   "TT426_5S_ALM_ANALOG_DB_VERY HIGH LEVEL VALUE (HH)" : Real = PLC TT426_5S_ALM_ANALOG_DB."VERY HIGH LEVEL VALUE (HH)" AT %DB2082.DBD34, 1 s
   "TT426_5S_ALM_ANALOG_DB_VERY LOW LEVEL VALUE (LL)" : Real = PLC TT426_5S_ALM_ANALOG_DB."VERY LOW LEVEL VALUE (LL)" AT %DB2082.DBD22, 1 s
   "TT426_6P_ALM_ANALOG_DB_HIGH LEVEL VALUE (H)" : Real = PLC TT426_6P_ALM_ANALOG_DB."HIGH LEVEL VALUE (H)" AT %DB2083.DBD30, 1 s
   "TT426_6P_ALM_ANALOG_DB_LOW LEVEL VALUE (L)" : Real = PLC TT426_6P_ALM_ANALOG_DB."LOW LEVEL VALUE (L)" AT %DB2083.DBD26, 1 s
   "TT426_6P_ALM_ANALOG_DB_VERY HIGH LEVEL VALUE (HH)" : Real = PLC TT426_6P_ALM_ANALOG_DB."VERY HIGH LEVEL VALUE (HH)" AT %DB2083.DBD34, 1 s
   "TT426_6P_ALM_ANALOG_DB_VERY LOW LEVEL VALUE (LL)" : Real = PLC TT426_6P_ALM_ANALOG_DB."VERY LOW LEVEL VALUE (LL)" AT %DB2083.DBD22, 1 s
   "TT426_6S_ALM_ANALOG_DB_HIGH LEVEL VALUE (H)" : Real = PLC TT426_6S_ALM_ANALOG_DB."HIGH LEVEL VALUE (H)" AT %DB2085.DBD30, 1 s
   "TT426_6S_ALM_ANALOG_DB_LOW LEVEL VALUE (L)" : Real = PLC TT426_6S_ALM_ANALOG_DB."LOW LEVEL VALUE (L)" AT %DB2085.DBD26, 1 s
   "TT426_6S_ALM_ANALOG_DB_VERY HIGH LEVEL VALUE (HH)" : Real = PLC TT426_6S_ALM_ANALOG_DB."VERY HIGH LEVEL VALUE (HH)" AT %DB2085.DBD34, 1 s
   "TT426_6S_ALM_ANALOG_DB_VERY LOW LEVEL VALUE (LL)" : Real = PLC TT426_6S_ALM_ANALOG_DB."VERY LOW LEVEL VALUE (LL)" AT %DB2085.DBD22, 1 s
   "TT426_APT_ALM_ANALOG_DB_HIGH LEVEL VALUE (H)" : Real = PLC TT426_APT_ALM_ANALOG_DB."HIGH LEVEL VALUE (H)" AT %DB2087.DBD30, 1 s
   "TT426_APT_ALM_ANALOG_DB_LOW LEVEL VALUE (L)" : Real = PLC TT426_APT_ALM_ANALOG_DB."LOW LEVEL VALUE (L)" AT %DB2087.DBD26, 1 s
   "TT426_APT_ALM_ANALOG_DB_VERY HIGH LEVEL VALUE (HH)" : Real = PLC TT426_APT_ALM_ANALOG_DB."VERY HIGH LEVEL VALUE (HH)" AT %DB2087.DBD34, 1 s
   "TT426_APT_ALM_ANALOG_DB_VERY LOW LEVEL VALUE (LL)" : Real = PLC TT426_APT_ALM_ANALOG_DB."VERY LOW LEVEL VALUE (LL)" AT %DB2087.DBD22, 1 s
   "TT426_FPT_ALM_ANALOG_DB_HIGH LEVEL VALUE (H)" : Real = PLC TT426_FPT_ALM_ANALOG_DB."HIGH LEVEL VALUE (H)" AT %DB2074.DBD30, 1 s
   "TT426_FPT_ALM_ANALOG_DB_LOW LEVEL VALUE (L)" : Real = PLC TT426_FPT_ALM_ANALOG_DB."LOW LEVEL VALUE (L)" AT %DB2074.DBD26, 1 s
   "TT426_FPT_ALM_ANALOG_DB_VERY HIGH LEVEL VALUE (HH)" : Real = PLC TT426_FPT_ALM_ANALOG_DB."VERY HIGH LEVEL VALUE (HH)" AT %DB2074.DBD34, 1 s
   "TT426_FPT_ALM_ANALOG_DB_VERY LOW LEVEL VALUE (LL)" : Real = PLC TT426_FPT_ALM_ANALOG_DB."VERY LOW LEVEL VALUE (LL)" AT %DB2074.DBD22, 1 s
   "TT426PORT_ALM_ANALOG_DB_HIGH LEVEL VALUE (H)" : Real = PLC TT426PORT_ALM_ANALOG_DB."HIGH LEVEL VALUE (H)" AT %DB2071.DBD30, 1 s
   "TT426PORT_ALM_ANALOG_DB_LOW LEVEL VALUE (L)" : Real = PLC TT426PORT_ALM_ANALOG_DB."LOW LEVEL VALUE (L)" AT %DB2071.DBD26, 1 s
   "TT426PORT_ALM_ANALOG_DB_VERY HIGH LEVEL VALUE (HH)" : Real = PLC TT426PORT_ALM_ANALOG_DB."VERY HIGH LEVEL VALUE (HH)" AT %DB2071.DBD34, 1 s
   "TT426PORT_ALM_ANALOG_DB_VERY LOW LEVEL VALUE (LL)" : Real = PLC TT426PORT_ALM_ANALOG_DB."VERY LOW LEVEL VALUE (LL)" AT %DB2071.DBD22, 1 s
   "TT426STR_ALM_ANALOG_DB_HIGH LEVEL VALUE (H)" : Real = PLC TT426STR_ALM_ANALOG_DB."HIGH LEVEL VALUE (H)" AT %DB2072.DBD30, 1 s
   "TT426STR_ALM_ANALOG_DB_LOW LEVEL VALUE (L)" : Real = PLC TT426STR_ALM_ANALOG_DB."LOW LEVEL VALUE (L)" AT %DB2072.DBD26, 1 s
   "TT426STR_ALM_ANALOG_DB_VERY HIGH LEVEL VALUE (HH)" : Real = PLC TT426STR_ALM_ANALOG_DB."VERY HIGH LEVEL VALUE (HH)" AT %DB2072.DBD34, 1 s
   "TT426STR_ALM_ANALOG_DB_VERY LOW LEVEL VALUE (LL)" : Real = PLC TT426STR_ALM_ANALOG_DB."VERY LOW LEVEL VALUE (LL)" AT %DB2072.DBD22, 1 s
   "LT421 1S  TANK LEVEL ALARM_ALARM L" : Bool = PLC "LT421 1S  TANK LEVEL ALARM"."ALARM L" AT %DB2228.DBX48.2, 1 s
   "LT421 2S  TANK LEVEL ALARM_ALARM L" : Bool = PLC "LT421 2S  TANK LEVEL ALARM"."ALARM L" AT %DB2230.DBX48.2, 1 s
   "LT421 3S  TANK LEVEL ALARM_ALARM L" : Bool = PLC "LT421 3S  TANK LEVEL ALARM"."ALARM L" AT %DB2232.DBX48.2, 1 s
   "LT421 4S  TANK LEVEL ALARM_ALARM L" : Bool = PLC "LT421 4S  TANK LEVEL ALARM"."ALARM L" AT %DB2234.DBX48.2, 1 s
   "LT421 5S  TANK LEVEL ALARM_ALARM L" : Bool = PLC "LT421 5S  TANK LEVEL ALARM"."ALARM L" AT %DB2236.DBX48.2, 1 s
   "LT421 6S  TANK LEVEL ALARM_ALARM L" : Bool = PLC "LT421 6S  TANK LEVEL ALARM"."ALARM L" AT %DB2238.DBX48.2, 1 s
   "LT422 1P  TANK LEVEL ALARM_ALARM L" : Bool = PLC "LT422 1P  TANK LEVEL ALARM"."ALARM L" AT %DB2227.DBX48.2, 1 s
   "LT422 3P  TANK LEVEL ALARM_ALARM L" : Bool = PLC "LT422 3P  TANK LEVEL ALARM"."ALARM L" AT %DB2231.DBX48.2, 1 s
   "LT422 4P  TANK LEVEL ALARM_ALARM L" : Bool = PLC "LT422 4P  TANK LEVEL ALARM"."ALARM L" AT %DB2233.DBX48.2, 1 s
   "LT422 4P  TANK LEVEL ALARM_HIGH LEVEL VALUE (H)" : Real = PLC "LT422 4P  TANK LEVEL ALARM"."HIGH LEVEL VALUE (H)" AT %DB2233.DBD30, 1 s
   "LT422 4P  TANK LEVEL ALARM_LOW LEVEL VALUE (L)" : Real = PLC "LT422 4P  TANK LEVEL ALARM"."LOW LEVEL VALUE (L)" AT %DB2233.DBD26, 1 s
   "LT422 4P  TANK LEVEL ALARM_VERY HIGH LEVEL VALUE (HH)" : Real = PLC "LT422 4P  TANK LEVEL ALARM"."VERY HIGH LEVEL VALUE (HH)" AT %DB2233.DBD34, 1 s
   "LT422 4P  TANK LEVEL ALARM_VERY LOW LEVEL VALUE (LL)" : Real = PLC "LT422 4P  TANK LEVEL ALARM"."VERY LOW LEVEL VALUE (LL)" AT %DB2233.DBD22, 1 s
   "LT422 5P  TANK LEVEL ALARM_ALARM L" : Bool = PLC "LT422 5P  TANK LEVEL ALARM"."ALARM L" AT %DB2235.DBX48.2, 1 s
   "LT422 6P  TANK LEVEL ALARM_ALARM L" : Bool = PLC "LT422 6P  TANK LEVEL ALARM"."ALARM L" AT %DB2237.DBX48.2, 1 s
   "LT422 APT  TANK LEVEL ALARM_ALARM L" : Bool = PLC "LT422 APT  TANK LEVEL ALARM"."ALARM L" AT %DB2239.DBX48.2, 1 s
   "LT422 FPT  TANK LEVEL ALARM_ALARM L" : Bool = PLC "LT422 FPT  TANK LEVEL ALARM"."ALARM L" AT %DB2226.DBX48.2, 1 s
   "LT422 FPT  TANK LEVEL ALARM_LOW LEVEL VALUE (L)" : Real = PLC "LT422 FPT  TANK LEVEL ALARM"."LOW LEVEL VALUE (L)" AT %DB2226.DBD26, 1 s
   "2084_Setpoints_Conf O2 Level Lo" : Real = PLC "2084_Setpoints"."Conf O2 Level Lo", 1 s
   "2084_Setpoints_Conf O2 Level Lo Lo" : Real = PLC "2084_Setpoints"."Conf O2 Level Lo Lo", 1 s
   "2084_Setpoints_DO_SP" : Real = PLC "2084_Setpoints".DO_SP AT %DB1.DBW0, 1 s
   "2084_Setpoints_FIT417_Hi" : Real = PLC "2084_Setpoints".FIT417_Hi, 1 s
   "2084_Setpoints_FIT417_HiHi" : Real = PLC "2084_Setpoints".FIT417_HiHi, 1 s
   "2084_Setpoints_FIT417_Lo" : Real = PLC "2084_Setpoints".FIT417_Lo, 1 s
   "2084_Setpoints_FIT417_LoLo" : Real = PLC "2084_Setpoints".FIT417_LoLo, 1 s
   "2084_Setpoints_FIT418_Hi" : Real = PLC "2084_Setpoints".FIT418_Hi AT %DB1.DBW0, 1 s
   "2084_Setpoints_FIT418_HiHi" : Real = PLC "2084_Setpoints".FIT418_HiHi AT %DB1.DBW0, 1 s
   "2084_Setpoints_FIT418_Lo" : Real = PLC "2084_Setpoints".FIT418_Lo AT %DB1.DBW0, 1 s
   "2084_Setpoints_FIT418_LoLo" : Real = PLC "2084_Setpoints".FIT418_LoLo AT %DB1.DBW0, 1 s
   "2084_Setpoints_FIT419_Hi" : Real = PLC "2084_Setpoints".FIT419_Hi, 1 s
   "2084_Setpoints_FIT419_HiHi" : Real = PLC "2084_Setpoints".FIT419_HiHi, 1 s
   "2084_Setpoints_FIT419_Lo" : Real = PLC "2084_Setpoints".FIT419_Lo, 1 s
   "2084_Setpoints_FIT419_LoLo" : Real = PLC "2084_Setpoints".FIT419_LoLo, 1 s
   "2084_Setpoints_FIT420_Hi" : Real = PLC "2084_Setpoints".FIT420_Hi AT %DB1.DBW0, 1 s
   "2084_Setpoints_FIT420_HiHi" : Real = PLC "2084_Setpoints".FIT420_HiHi AT %DB1.DBW0, 1 s
   "2084_Setpoints_FIT420_Lo" : Real = PLC "2084_Setpoints".FIT420_Lo AT %DB1.DBW0, 1 s
   "2084_Setpoints_FIT420_LoLo" : Real = PLC "2084_Setpoints".FIT420_LoLo AT %DB1.DBW0, 1 s
   "2084_Setpoints_LT421_Hi" : Real = PLC "2084_Setpoints".LT421_Hi, 1 s
   "2084_Setpoints_LT421_Lo" : Real = PLC "2084_Setpoints".LT421_Lo, 1 s
   "2084_Setpoints_LT422_Hi" : Real = PLC "2084_Setpoints".LT422_Hi AT %DB1.DBW0, 1 s
   "2084_Setpoints_LT422_Lo" : Real = PLC "2084_Setpoints".LT422_Lo AT %DB1.DBW0, 1 s
   "2084_Setpoints_PH_SP" : Real = PLC "2084_Setpoints".PH_SP AT %DB1.DBW0, 1 s
   "2084_Setpoints_PIT415_Hi" : Real = PLC "2084_Setpoints".PIT415_Hi AT %DB1.DBW0, 1 s
   "2084_Setpoints_PIT415_HiHi" : Real = PLC "2084_Setpoints".PIT415_HiHi AT %DB1.DBW0, 1 s
   "2084_Setpoints_PIT415_Lo" : Real = PLC "2084_Setpoints".PIT415_Lo AT %DB1.DBW0, 1 s
   "2084_Setpoints_PIT415_LoLo" : Real = PLC "2084_Setpoints".PIT415_LoLo AT %DB1.DBW0, 1 s
   "2084_Setpoints_PIT424_Hi" : Real = PLC "2084_Setpoints".PIT424_Hi AT %DB1.DBW0, 1 s
   "2084_Setpoints_PIT424_HiHi" : Real = PLC "2084_Setpoints".PIT424_HiHi AT %DB1.DBW0, 1 s
   "2084_Setpoints_PIT424_Lo" : Real = PLC "2084_Setpoints".PIT424_Lo AT %DB1.DBW0, 1 s
   "2084_Setpoints_PIT424_LoLo" : Real = PLC "2084_Setpoints".PIT424_LoLo AT %DB1.DBW0, 1 s
   "2084_Setpoints_TT436_Hi" : Real = PLC "2084_Setpoints".TT436_Hi AT %DB1.DBW0, 1 s
   "2084_Setpoints_TT436_HiHi" : Real = PLC "2084_Setpoints".TT436_HiHi AT %DB1.DBW0, 1 s
   "2084_Setpoints_TX426 PH High" : Real = PLC "2084_Setpoints"."TX426 Port PH High", 1 s
   "2084_Setpoints_TX426 PH Lo" : Real = PLC "2084_Setpoints"."TX426 Port PH Lo", 1 s
   "2084_Setpoints_TX426 Star PH High" : Real = PLC "2084_Setpoints"."TX425 Star PH High", 1 s
   "2084_Setpoints_TX426 Star PH Lo" : Real = PLC "2084_Setpoints"."TX425 Star PH Lo", 1 s
   "2084_Setpoints_TX428 DO High" : Real = PLC "2084_Setpoints"."TX428 Port DO High", 1 s
   "2084_Setpoints_TX428 DO Lo" : Real = PLC "2084_Setpoints"."TX428 Port DO Lo", 1 s
   "2084_Setpoints_TX428 Star DO High" : Real = PLC "2084_Setpoints"."TX427 Star DO High", 1 s
   "2084_Setpoints_TX428 Star DO Lo" : Real = PLC "2084_Setpoints"."TX427 Star DO Lo", 1 s
   "BRIGE HMI HEART BEAT" : Bool = PLC "59_COMMS_HEALTH_DATA"."BRIGE HMI HB" AT %DB1.DBX0.0, 100 ms
   "TRUE" : Bool = PLC AlwaysTRUE AT %M1.2, 1 s
   "IGG PLC HEART BEAT" : Bool = PLC "55_STATUS_DATA".HEART_BEAT AT %DB55.DBX0.0, 100 ms
      on ChangeValue: "HeartBeatFunction"()
   "Setpoint Override_DB_Set Pressure" : Bool = PLC "Setpoint Override_DB"."Set Pressure", 1 s
   "Warn To Start IGG" : Bool = PLC "82_To_HMI"."Warn to Start IGG", 1 s
      on ChangeValue: "TreatmentRequired"()
   "Warn To Start IGG-Last" : Bool = PLC "82_To_HMI"."Warn to Start IGG-Last", 1 s
      on ChangeValue: "TimeRemainingToTreatment"()
   "Warn To Start GCU" : Bool = PLC "82_To_HMI"."Warn to Start GCU", 1 s
      on ChangeValue: "TimeRemainingToRe_Ox"()
   "Warn To Start GCU-Last" : Bool = PLC "82_To_HMI"."Warn to Start GCU-Last", 1 s

discrete alarms
   33: 'TIT-315 SHELL CSW TEMP - HIGH HIGH AND FS-317 - FAULT', class IGG Alarms, trigger "Alarms_Acknowledge_IGG_ALARM_ACKNLG_3" bit 0
   34: 'TIT-315 SHELL CSW TEMP - HIGH HIGH AND TS-006 - FAULT', class IGG Alarms, trigger "Alarms_Acknowledge_IGG_ALARM_ACKNLG_3" bit 1
   35: 'TIT-315 SHELL CSW TEMP - HIGH HIGH AND TIT-401 - FAULT', class IGG Alarms, trigger "Alarms_Acknowledge_IGG_ALARM_ACKNLG_3" bit 2
   36: 'PIT-316 OUTLET CSW PRESSURE AND FS-317 - FAULT', class IGG Alarms, trigger "Alarms_Acknowledge_IGG_ALARM_ACKNLG_3" bit 3
   37: 'PIT-316 OUTLET CSW PRESSURE AND TIT-315 - FAULT', class IGG Alarms, trigger "Alarms_Acknowledge_IGG_ALARM_ACKNLG_3" bit 4
   38: 'PIT-316 OUTLET CSW PRESSURE AND TS-006 - FAULT', class IGG Alarms, trigger "Alarms_Acknowledge_IGG_ALARM_ACKNLG_3" bit 5
   39: 'IGG_ALARM_WORD_03_BIT_14', class IGG Alarms, trigger "Alarms_Acknowledge_IGG_ALARM_ACKNLG_3" bit 6
   40: 'IGG_ALARM_WORD_03_BIT_15', class IGG Alarms, trigger "Alarms_Acknowledge_IGG_ALARM_ACKNLG_3" bit 7
   41: 'PIT-112/113 TIER ALARM - PRESSURE NOT OK', class IGG Alarms, trigger "Alarms_Acknowledge_IGG_ALARM_ACKNLG_3" bit 8
   42: 'PIT-102 CA PRESSURE - LOW LOW AND FDU - FAULT', class IGG Alarms, trigger "Alarms_Acknowledge_IGG_ALARM_ACKNLG_3" bit 9
   43: 'PIT-102 CA PRESSURE - LOW LOW AND PIT-402 - FAULT', class IGG Alarms, trigger "Alarms_Acknowledge_IGG_ALARM_ACKNLG_3" bit 10
   44: 'IGG ALARM WORD', class IGG Alarms, trigger "Alarms_Acknowledge_IGG_ALARM_ACKNLG_3" bit 11
   45: 'TIT-401 IG TEMP - HIGH HIGH AND TS-403 - FAULT', class IGG Alarms, trigger "Alarms_Acknowledge_IGG_ALARM_ACKNLG_3" bit 12
   46: 'TIT-401 IG TEMP - HIGH HIGH AND TIT-360 - FAULT', class IGG Alarms, trigger "Alarms_Acknowledge_IGG_ALARM_ACKNLG_3" bit 13
   47: 'IGG_ALARM_WORD_03_BIT_6', class IGG Alarms, trigger "Alarms_Acknowledge_IGG_ALARM_ACKNLG_3" bit 14
   48: 'IGG_ALARM_WORD_03_BIT_7', class IGG Alarms, trigger "Alarms_Acknowledge_IGG_ALARM_ACKNLG_3" bit 15
   49: 'TIT-319 INLET CSW TEMP - FAULT AND TS-006 - FAULT', class IGG Alarms, trigger "Alarms_Acknowledge_IGG_ALARM_ACKNLG_4" bit 0
   50: 'TIT-319 INLET CSW TEMP - FAULT AND TIT-401 AND TIT-360 - FAULT', class IGG Alarms, trigger "Alarms_Acknowledge_IGG_ALARM_ACKNLG_4" bit 1
   51: 'TIT-360 OUTLET CSW TEMP - HIGH HIGH0', class IGG Alarms, trigger "Alarms_Acknowledge_IGG_ALARM_ACKNLG_4" bit 2
   52: 'TIT-360 OUTLET CSW TEMP - HIGH HIGH AND TIT-401 - FAULT', class IGG Alarms, trigger "Alarms_Acknowledge_IGG_ALARM_ACKNLG_4" bit 3
   53: 'E-139 NOT RUNNING2', class IGG Alarms, trigger "Alarms_Acknowledge_IGG_ALARM_ACKNLG_4" bit 4
   54: 'CORRECT PHASE ROTATION - FAULT', class IGG Alarms, trigger "Alarms_Acknowledge_IGG_ALARM_ACKNLG_4" bit 5
   55: 'IGG_ALARM_WORD_04_BIT_14', class IGG Alarms, trigger "Alarms_Acknowledge_IGG_ALARM_ACKNLG_4" bit 6
   56: 'IGG_ALARM_WORD_04_BIT_15', class IGG Alarms, trigger "Alarms_Acknowledge_IGG_ALARM_ACKNLG_4" bit 7
   57: 'CV-311 - FAULT', class IGG Alarms, trigger "Alarms_Acknowledge_IGG_ALARM_ACKNLG_4" bit 8
   58: 'CV-312 - FAULT', class IGG Alarms, trigger "Alarms_Acknowledge_IGG_ALARM_ACKNLG_4" bit 9
   59: 'CV-321 - FAULT', class IGG Alarms, trigger "Alarms_Acknowledge_IGG_ALARM_ACKNLG_4" bit 10
   60: 'CV-322 - FAULT', class IGG Alarms, trigger "Alarms_Acknowledge_IGG_ALARM_ACKNLG_4" bit 11
   61: 'CV-401 - FAULT', class IGG Alarms, trigger "Alarms_Acknowledge_IGG_ALARM_ACKNLG_4" bit 12
   62: 'CV-431 - FAULT', class IGG Alarms, trigger "Alarms_Acknowledge_IGG_ALARM_ACKNLG_4" bit 13
   63: 'CV-432 - FAULT', class IGG Alarms, trigger "Alarms_Acknowledge_IGG_ALARM_ACKNLG_4" bit 14
   64: 'SAFETY SYSTEM INTERLOCK', class IGG Alarms, trigger "Alarms_Acknowledge_IGG_ALARM_ACKNLG_4" bit 15
   65: 'IGG ALARM ACTIVE', class BC Alarms, trigger "BC_ALARM_ACKNLG_1" bit 0
   66: 'PS-101 PRESSURE NOT PRESENT - FAULT', class BC Alarms, trigger "BC_ALARM_ACKNLG_1" bit 1
   67: 'E-600 O2 ANALYSER SYSTEM - FAIL', class BC Alarms, trigger "BC_ALARM_ACKNLG_1" bit 2
   68: 'O2 SYSTEM POWER NOT HEALTHY', class BC Alarms, trigger "BC_ALARM_ACKNLG_1" bit 3
   69: 'FD-001 FLAME SIGNAL - OUT OF RANGE', class BC Alarms, trigger "BC_ALARM_ACKNLG_1" bit 4
   70: 'E-600 O2 ANALYSER CONTENT - OUT OF RANGE', class BC Alarms, trigger "BC_ALARM_ACKNLG_1" bit 5
   71: 'E-600 O2 ANALYSER CONTENT - LOW LOW', class BC Alarms, trigger "BC_ALARM_ACKNLG_1" bit 6
   72: 'BC_ALARM_WORD_01_BIT_15', class BC Alarms, trigger "BC_ALARM_ACKNLG_1" bit 7
   73: 'MASTER PLC HEART BEAT MISSING', class BC Alarms, trigger "BC_ALARM_ACKNLG_1" bit 8
   74: 'IGNITER POWER NOT HEALTHY', class BC Alarms, trigger "BC_ALARM_ACKNLG_1" bit 9
   75: 'BC AUTO INTERLOCKS NOT OK', class BC Alarms, trigger "BC_ALARM_ACKNLG_1" bit 10
   76: 'FDU POWER NOT HEALTHY', class BC Alarms, trigger "BC_ALARM_ACKNLG_1" bit 11
   77: 'PILOT FLAME IGNITION SEQUENCE FAILURE', class BC Alarms, trigger "BC_ALARM_ACKNLG_1" bit 12
   78: 'MAIN BURNER FLAME SEQUENCE FAILURE', class BC Alarms, trigger "BC_ALARM_ACKNLG_1" bit 13
   79: 'PILOT FLAME PURGE SEQUENCE FAILURE', class BC Alarms, trigger "BC_ALARM_ACKNLG_1" bit 14
   80: 'FD-001 FLAME DETECTION UNIT NOT HEALTHY', class BC Alarms, trigger "BC_ALARM_ACKNLG_1" bit 15
   81: 'PIT-204 FUEL OIL INLET PRESSURE READING - FAULT AND PIT-205 - FAULT', class BC Alarms, trigger "BC_ALARM_ACKNLG_2" bit 0
   82: 'PIT-204 FUEL OIL INLET PRESSURE READING - FAULT AND CV-206 AND CV-207 - CLOSED', class BC Alarms, trigger "BC_ALARM_ACKNLG_2" bit 1
   83: 'BC_ALARM_WORD_02_BIT_10', class BC Alarms, trigger "BC_ALARM_ACKNLG_2" bit 2
   84: 'PIT-204 FUEL OIL INLET PRESSURE LOW LOW AND PIT-205 - FAULT', class BC Alarms, trigger "BC_ALARM_ACKNLG_2" bit 3
   85: 'PIT-204 FUEL OIL INLET PRESSURE - LOW LOW', class BC Alarms, trigger "BC_ALARM_ACKNLG_2" bit 4
   86: 'PIT-204 FUEL OIL INLET PRESSURE - HIGH HIGH AND PIT-205 - FAULT', class BC Alarms, trigger "BC_ALARM_ACKNLG_2" bit 5
   87: 'PIT-204 FUEL OIL INLET PRESSURE - HIGH HIGH AND CV-206 AND CV-207 CLOSED', class BC Alarms, trigger "BC_ALARM_ACKNLG_2" bit 6
   88: 'BC_ALARM_WORD_02_BIT_15', class BC Alarms, trigger "BC_ALARM_ACKNLG_2" bit 7
   89: 'NO FLOW AT FS-317', class BC Alarms, trigger "BC_ALARM_ACKNLG_2" bit 8
   90: 'NO FLOW AT FS-320', class BC Alarms, trigger "BC_ALARM_ACKNLG_2" bit 9
   91: 'BC_ALARM_WORD_02_BIT_2', class BC Alarms, trigger "BC_ALARM_ACKNLG_2" bit 10
   92: 'BC_ALARM_WORD_02_BIT_3', class BC Alarms, trigger "BC_ALARM_ACKNLG_2" bit 11
   93: 'BC_ALARM_WORD_02_BIT_4', class BC Alarms, trigger "BC_ALARM_ACKNLG_2" bit 12
   94: 'BC_ALARM_WORD_02_BIT_5', class BC Alarms, trigger "BC_ALARM_ACKNLG_2" bit 13
   95: 'BC_ALARM_WORD_02_BIT_6', class BC Alarms, trigger "BC_ALARM_ACKNLG_2" bit 14
   96: 'BC_ALARM_WORD_02_BIT_7', class BC Alarms, trigger "BC_ALARM_ACKNLG_2" bit 15
   97: 'FS-320 COOLING WATER FLOW SWITCH - FAULT AND FS-317 - FAULT', class BC Alarms, trigger "BC_ALARM_ACKNLG_3" bit 0
   98: 'FS-320 COOLING WATER FLOW SWITCH - FAULT AND TIT-360 - FAULT', class BC Alarms, trigger "BC_ALARM_ACKNLG_3" bit 1
   99: 'FS-320 COOLING WATER FLOW SWITCH - FAULT AND TIT-401 - FAULT0', class BC Alarms, trigger "BC_ALARM_ACKNLG_3" bit 2
   100: 'FS-317 JACKET COOLING WATER FLOW SWITCH - FAULT AND FS-320 - FAULT AND PIT 360 - FAULT', class BC Alarms, trigger "BC_ALARM_ACKNLG_3" bit 3
   101: 'FS-317 JACKET COOLING WATER FLOW SWITCH FASULT AND TIT-360 - FAULT', class BC Alarms, trigger "BC_ALARM_ACKNLG_3" bit 4
   102: 'FS-317 JACKET COOLING WATER FLOW SWITCH - FAULT AND TIT-401 - FAULT', class BC Alarms, trigger "BC_ALARM_ACKNLG_3" bit 5
   103: 'BC_ALARM_WORD_03_BIT_14', class BC Alarms, trigger "BC_ALARM_ACKNLG_3" bit 6
   104: 'TS-403 IG VENT TEMPERATURE HIGH', class BC Alarms, trigger "BC_ALARM_ACKNLG_3" bit 7
   105: 'FS-123 PILOT BURNER AIR FLOW SWITCH - FAULT AND PIT-112 HIGH HIGH', class BC Alarms, trigger "BC_ALARM_ACKNLG_3" bit 8
   106: 'FS-123 PILOT BURNER AIR FLOW SWITCH - FAULT AND PIT-112 LOW LOW', class BC Alarms, trigger "BC_ALARM_ACKNLG_3" bit 9
   107: 'PIT-112 INSTRUMENT AIR PRESSURE - FAULT', class BC Alarms, trigger "BC_ALARM_ACKNLG_3" bit 10
   108: 'PIT-112 INSTRUMENT AIR PRESSURE - FAULT AND FS-115 - FAULT', class BC Alarms, trigger "BC_ALARM_ACKNLG_3" bit 11
   109: 'FS-115 MAIN BURNER ATOMISING AIR FLOW SWITCH - FAULT AND CV 114 CLOSE', class BC Alarms, trigger "BC_ALARM_ACKNLG_3" bit 12
   110: 'FS-115 MAIN BURNER ATOMISING AIR FLOW SWITCH - FAULT AND PIT-113 - FAULT', class BC Alarms, trigger "BC_ALARM_ACKNLG_3" bit 13
   111: 'BC_ALARM_WORD_03_BIT_6', class BC Alarms, trigger "BC_ALARM_ACKNLG_3" bit 14
   112: 'BC_ALARM_WORD_3_BIT_15', class BC Alarms, trigger "BC_ALARM_ACKNLG_3" bit 15
   113: 'LS-001 IGG QUENCH CHAMBER LEVEL - HIGH', class BC Alarms, trigger "BC_ALARM_ACKNLG_4" bit 0
   114: 'P-305 FRESH WATER PUMP - TRIPPED', class BC Alarms, trigger "BC_ALARM_ACKNLG_4" bit 1
   115: 'BC_ALARM_WORD_04_BIT_10', class BC Alarms, trigger "BC_ALARM_ACKNLG_4" bit 2
   116: 'BC_ALARM_WORD_04_BIT_11', class BC Alarms, trigger "BC_ALARM_ACKNLG_4" bit 3
   117: 'BC_ALARM_WORD_04_BIT_12', class BC Alarms, trigger "BC_ALARM_ACKNLG_4" bit 4
   118: 'BC_ALARM_WORD_04_BIT_13', class BC Alarms, trigger "BC_ALARM_ACKNLG_4" bit 5
   119: 'BC_ALARM_WORD_04_BIT_14', class BC Alarms, trigger "BC_ALARM_ACKNLG_4" bit 6
   120: 'BC_ALARM_WORD_04_BIT_15', class BC Alarms, trigger "BC_ALARM_ACKNLG_4" bit 7
   121: 'TS-006 IGG SHELL TEMPERATURE - HIGH', class BC Alarms, trigger "BC_ALARM_ACKNLG_4" bit 8
   122: 'TS-006 IG SHELL TEMP HI SWITCH AND TIT-360 - FAULT', class BC Alarms, trigger "BC_ALARM_ACKNLG_4" bit 9
   123: 'TS-006 IG SHELL TEMP HI SWITCH AND TIT-401 - FAULT', class BC Alarms, trigger "BC_ALARM_ACKNLG_4" bit 10
   124: 'TS-403 IG TEMP - HIGH HIGH SWITCH AND TIT-401 - FAULT', class BC Alarms, trigger "BC_ALARM_ACKNLG_4" bit 11
   125: 'TS-403 IG TEMP - HIGH HIGH SWITCH AND TIT-360 - FAULT', class BC Alarms, trigger "BC_ALARM_ACKNLG_4" bit 12
   126: 'PIT-113 IGG MAIN ATOM AIR PRESSURE - FAULT', class BC Alarms, trigger "BC_ALARM_ACKNLG_4" bit 13
   127: 'PIT-205 IGG MAIN FUEL PRESSURE - FAULT', class BC Alarms, trigger "BC_ALARM_ACKNLG_4" bit 14
   128: 'TIT-202 IGG INLET FUEL TEMP', class BC Alarms, trigger "BC_ALARM_ACKNLG_4" bit 15
   129: 'PIT-359 - HIGH HIGH', class IGG Alarms, trigger "Alarms_Acknowledge_IGG_ALARM_ACKNLG_2" bit 1
   130: 'PIT-316 - HIGH HIGH', class IGG Alarms, trigger "Alarms_Acknowledge_IGG_ALARM_ACKNLG_2" bit 3
   131: 'PIT-359 - LOW LOW', class IGG Alarms, trigger "Alarms_Acknowledge_IGG_ALARM_ACKNLG_2" bit 0
   132: 'PIT-316 - LOW LOW', class IGG Alarms, trigger "Alarms_Acknowledge_IGG_ALARM_ACKNLG_2" bit 2
   133: 'PIT-359 - HIGH HIGH', class IGG Alarms, trigger "Alarms_Acknowledge_IGG_ALARM_ACKNLG_2" bit 4
   134: 'TIT-401 - HIGH HIGH', class IGG Alarms, trigger "Alarms_Acknowledge_IGG_ALARM_ACKNLG_2" bit 10
   135: 'PIT-102 CA PRESSURE - FAULT', class IGG Alarms, trigger "Alarms_Acknowledge_IGG_ALARM_ACKNLG_2" bit 9
   136: 'PIT-402 IG OUTLET PRESSURE - HIGH HIGH', class IGG Alarms, trigger "Alarms_Acknowledge_IGG_ALARM_ACKNLG_2" bit 12
   137: 'PIT-402 IG OUTLET PRESSURE - LOW LOW', class IGG Alarms, trigger "Alarms_Acknowledge_IGG_ALARM_ACKNLG_2" bit 11
   138: 'IGG_ALARM_WORD_02_BIT_14', class IGG Alarms, trigger "Alarms_Acknowledge_IGG_ALARM_ACKNLG_2" bit 6
   139: 'IGG_ALARM_WORD_02_BIT_13', class IGG Alarms, trigger "Alarms_Acknowledge_IGG_ALARM_ACKNLG_2" bit 5
   140: 'PIT-102 CA PRESSURE - LOW LOW', class IGG Alarms, trigger "Alarms_Acknowledge_IGG_ALARM_ACKNLG_2" bit 8
   141: 'IGG_ALARM_WORD_02_BIT_15', class IGG Alarms, trigger "Alarms_Acknowledge_IGG_ALARM_ACKNLG_2" bit 7
   142: 'EMERGENCY STOP ACTIVE', class IGG Alarms, trigger "Alarms_Acknowledge_IGG_ALARM_ACKNLG_1" bit 15
   143: 'ATMOSPHERIC O2 SENSOR 1 - LOW LOW', class IGG Alarms, trigger "Alarms_Acknowledge_IGG_ALARM_ACKNLG_1" bit 1
   144: 'BC ALARM ACTIVE', class IGG Alarms, trigger "Alarms_Acknowledge_IGG_ALARM_ACKNLG_1" bit 0
   145: 'ATMOSPHERIC O2 SENSOR 2 - LOW LOW', class IGG Alarms, trigger "Alarms_Acknowledge_IGG_ALARM_ACKNLG_1" bit 2
   146: 'E-500B FUEL PUMP - NOT RUNNING', class IGG Alarms, trigger "Alarms_Acknowledge_IGG_ALARM_ACKNLG_1" bit 4
   147: 'E-500A FUEL PUMP - NOT RUNNING', class IGG Alarms, trigger "Alarms_Acknowledge_IGG_ALARM_ACKNLG_1" bit 3
   148: 'P-301 CSW PUMP - TRIPPED', class IGG Alarms, trigger "Alarms_Acknowledge_IGG_ALARM_ACKNLG_1" bit 11
   149: 'IGG AUTO INTERLOCKS NOT OK', class IGG Alarms, trigger "Alarms_Acknowledge_IGG_ALARM_ACKNLG_1" bit 10
   150: 'E-500A FUEL PUMP - TRIPPED', class IGG Alarms, trigger "Alarms_Acknowledge_IGG_ALARM_ACKNLG_1" bit 12
   151: 'E-139 CAB INVERTER - FAULT', class IGG Alarms, trigger "Alarms_Acknowledge_IGG_ALARM_ACKNLG_1" bit 14
   152: 'E-500B FUEL PUMP - TRIPPED', class IGG Alarms, trigger "Alarms_Acknowledge_IGG_ALARM_ACKNLG_1" bit 13
   153: 'IGG_ALARM_WORD_01_BIT_14', class IGG Alarms, trigger "Alarms_Acknowledge_IGG_ALARM_ACKNLG_1" bit 6
   154: 'E-139 CAB NOT READY3', class IGG Alarms, trigger "Alarms_Acknowledge_IGG_ALARM_ACKNLG_1" bit 5
   155: 'IGG_ALARM_WORD_01_BIT_15', class IGG Alarms, trigger "Alarms_Acknowledge_IGG_ALARM_ACKNLG_1" bit 7
   156: 'SLAVE PLC HEART BEAT MISSING', class IGG Alarms, trigger "Alarms_Acknowledge_IGG_ALARM_ACKNLG_1" bit 9
   157: 'MASTER PLC HEART BEAT MISSING', class IGG Alarms, trigger "Alarms_Acknowledge_IGG_ALARM_ACKNLG_1" bit 8
   158: 'PIT-402 IG PRESSURE - OUT OF RANGE', class IGG Alarms, trigger "Alarms_Acknowledge_IGG_ALARM_ACKNLG_2" bit 13
   159: 'TIT-360 - HIGH HIGH', class IGG Alarms, trigger "Alarms_Acknowledge_IGG_ALARM_ACKNLG_2" bit 15
   160: 'TIT-319 - HIGH HIGH', class IGG Alarms, trigger "Alarms_Acknowledge_IGG_ALARM_ACKNLG_2" bit 14
   257: 'IGG_MESSAGE_WORD_01_BIT_8', class IGG Messages, trigger "64_Message_Data_IGG_MESSAGE_WORD_01" bit 0
   258: 'IGG_MESSAGE_WORD_01_BIT_9', class IGG Messages, trigger "64_Message_Data_IGG_MESSAGE_WORD_01" bit 1
   259: 'IGG_MESSAGE_WORD_01_BIT_10', class IGG Messages, trigger "64_Message_Data_IGG_MESSAGE_WORD_01" bit 2
   260: 'IGG_MESSAGE_WORD_01_BIT_11', class IGG Messages, trigger "64_Message_Data_IGG_MESSAGE_WORD_01" bit 3
   261: 'IGG_MESSAGE_WORD_01_BIT_12', class IGG Messages, trigger "64_Message_Data_IGG_MESSAGE_WORD_01" bit 4
   262: 'IGG_MESSAGE_WORD_01_BIT_13', class IGG Messages, trigger "64_Message_Data_IGG_MESSAGE_WORD_01" bit 5
   263: 'IGG_MESSAGE_WORD_01_BIT_14', class IGG Messages, trigger "64_Message_Data_IGG_MESSAGE_WORD_01" bit 6
   264: 'IGG_MESSAGE_WORD_01_BIT_15', class IGG Messages, trigger "64_Message_Data_IGG_MESSAGE_WORD_01" bit 7
   265: 'IGG_MESSAGE_WORD_01_BIT_0', class IGG Messages, trigger "64_Message_Data_IGG_MESSAGE_WORD_01" bit 8
   266: 'IGG_MESSAGE_WORD_01_BIT_1', class IGG Messages, trigger "64_Message_Data_IGG_MESSAGE_WORD_01" bit 9
   267: 'IGG_MESSAGE_WORD_01_BIT_2', class IGG Messages, trigger "64_Message_Data_IGG_MESSAGE_WORD_01" bit 10
   268: 'IGG_MESSAGE_WORD_01_BIT_3', class IGG Messages, trigger "64_Message_Data_IGG_MESSAGE_WORD_01" bit 11
   269: 'IGG_MESSAGE_WORD_01_BIT_4', class IGG Messages, trigger "64_Message_Data_IGG_MESSAGE_WORD_01" bit 12
   270: 'IGG_MESSAGE_WORD_01_BIT_5', class IGG Messages, trigger "64_Message_Data_IGG_MESSAGE_WORD_01" bit 13
   271: 'IGG_MESSAGE_WORD_01_BIT_6', class IGG Messages, trigger "64_Message_Data_IGG_MESSAGE_WORD_01" bit 14
   272: 'IGG_MESSAGE_WORD_01_BIT_7', class IGG Messages, trigger "64_Message_Data_IGG_MESSAGE_WORD_01" bit 15
   273: 'IGG_MESSAGE_WORD_02_BIT_8', class IGG Messages, trigger "64_Message_Data_IGG_MESSAGE_WORD_02" bit 0
   274: 'IGG_MESSAGE_WORD_02_BIT_9', class IGG Messages, trigger "64_Message_Data_IGG_MESSAGE_WORD_02" bit 1
   275: 'IGG_MESSAGE_WORD_02_BIT_10', class IGG Messages, trigger "64_Message_Data_IGG_MESSAGE_WORD_02" bit 2
   276: 'IGG_MESSAGE_WORD_02_BIT_11', class IGG Messages, trigger "64_Message_Data_IGG_MESSAGE_WORD_02" bit 3
   277: 'IGG_MESSAGE_WORD_02_BIT_12', class IGG Messages, trigger "64_Message_Data_IGG_MESSAGE_WORD_02" bit 4
   278: 'IGG_MESSAGE_WORD_02_BIT_13', class IGG Messages, trigger "64_Message_Data_IGG_MESSAGE_WORD_02" bit 5
   279: 'IGG_MESSAGE_WORD_02_BIT_14', class IGG Messages, trigger "64_Message_Data_IGG_MESSAGE_WORD_02" bit 6
   280: 'IGG_MESSAGE_WORD_02_BIT_15', class IGG Messages, trigger "64_Message_Data_IGG_MESSAGE_WORD_02" bit 7
   281: 'IGG_MESSAGE_WORD_02_BIT_0', class IGG Messages, trigger "64_Message_Data_IGG_MESSAGE_WORD_02" bit 8
   282: 'IGG_MESSAGE_WORD_02_BIT_1', class IGG Messages, trigger "64_Message_Data_IGG_MESSAGE_WORD_02" bit 9
   283: 'IGG_MESSAGE_WORD_02_BIT_2', class IGG Messages, trigger "64_Message_Data_IGG_MESSAGE_WORD_02" bit 10
   284: 'IGG_MESSAGE_WORD_02_BIT_3', class IGG Messages, trigger "64_Message_Data_IGG_MESSAGE_WORD_02" bit 11
   285: 'IGG_MESSAGE_WORD_02_BIT_4', class IGG Messages, trigger "64_Message_Data_IGG_MESSAGE_WORD_02" bit 12
   286: 'IGG_MESSAGE_WORD_02_BIT_5', class IGG Messages, trigger "64_Message_Data_IGG_MESSAGE_WORD_02" bit 13
   287: 'IGG_MESSAGE_WORD_02_BIT_6', class IGG Messages, trigger "64_Message_Data_IGG_MESSAGE_WORD_02" bit 14
   288: 'IGG_MESSAGE_WORD_02_BIT_7', class IGG Messages, trigger "64_Message_Data_IGG_MESSAGE_WORD_02" bit 15
   289: 'BC_MESSAGE_WORD_01_BIT_8', class BC Messages, trigger "64_Message_Data_BC_MESSAGE_WORD_01" bit 0
   290: 'BC_MESSAGE_WORD_01_BIT_9', class BC Messages, trigger "64_Message_Data_BC_MESSAGE_WORD_01" bit 1
   291: 'BC_MESSAGE_WORD_01_BIT_10', class BC Messages, trigger "64_Message_Data_BC_MESSAGE_WORD_01" bit 2
   292: 'BC_MESSAGE_WORD_01_BIT_11', class BC Messages, trigger "64_Message_Data_BC_MESSAGE_WORD_01" bit 3
   293: 'BC_MESSAGE_WORD_01_BIT_12', class BC Messages, trigger "64_Message_Data_BC_MESSAGE_WORD_01" bit 4
   294: 'BC_MESSAGE_WORD_01_BIT_13', class BC Messages, trigger "64_Message_Data_BC_MESSAGE_WORD_01" bit 5
   295: 'BC_MESSAGE_WORD_01_BIT_14', class BC Messages, trigger "64_Message_Data_BC_MESSAGE_WORD_01" bit 6
   296: 'BC_MESSAGE_WORD_01_BIT_15', class BC Messages, trigger "64_Message_Data_BC_MESSAGE_WORD_01" bit 7
   297: 'BC_MESSAGE_WORD_01_BIT_0', class BC Messages, trigger "64_Message_Data_BC_MESSAGE_WORD_01" bit 8
   298: 'BC_MESSAGE_WORD_01_BIT_1', class BC Messages, trigger "64_Message_Data_BC_MESSAGE_WORD_01" bit 9
   299: 'BC_MESSAGE_WORD_01_BIT_2', class BC Messages, trigger "64_Message_Data_BC_MESSAGE_WORD_01" bit 10
   300: 'BC_MESSAGE_WORD_01_BIT_3', class BC Messages, trigger "64_Message_Data_BC_MESSAGE_WORD_01" bit 11
   301: 'BC_MESSAGE_WORD_01_BIT_4', class BC Messages, trigger "64_Message_Data_BC_MESSAGE_WORD_01" bit 12
   302: 'BC_MESSAGE_WORD_01_BIT_5', class BC Messages, trigger "64_Message_Data_BC_MESSAGE_WORD_01" bit 13
   303: 'BC_MESSAGE_WORD_01_BIT_6', class BC Messages, trigger "64_Message_Data_BC_MESSAGE_WORD_01" bit 14
   304: 'BC_MESSAGE_WORD_01_BIT_7', class BC Messages, trigger "64_Message_Data_BC_MESSAGE_WORD_01" bit 15
   305: 'BC_MESSAGE_WORD_02_BIT_8', class BC Messages, trigger "64_Message_Data_BC_MESSAGE_WORD_02" bit 0
   306: 'BC_MESSAGE_WORD_02_BIT_9', class BC Messages, trigger "64_Message_Data_BC_MESSAGE_WORD_02" bit 1
   307: 'BC_MESSAGE_WORD_02_BIT_10', class BC Messages, trigger "64_Message_Data_BC_MESSAGE_WORD_02" bit 2
   308: 'BC_MESSAGE_WORD_02_BIT_11', class BC Messages, trigger "64_Message_Data_BC_MESSAGE_WORD_02" bit 3
   309: 'BC_MESSAGE_WORD_02_BIT_12', class BC Messages, trigger "64_Message_Data_BC_MESSAGE_WORD_02" bit 4
   310: 'BC_MESSAGE_WORD_02_BIT_13', class BC Messages, trigger "64_Message_Data_BC_MESSAGE_WORD_02" bit 5
   311: 'BC_MESSAGE_WORD_02_BIT_14', class BC Messages, trigger "64_Message_Data_BC_MESSAGE_WORD_02" bit 6
   312: 'BC_MESSAGE_WORD_02_BIT_15', class BC Messages, trigger "64_Message_Data_BC_MESSAGE_WORD_02" bit 7
   313: 'BC_MESSAGE_WORD_02_BIT_0', class BC Messages, trigger "64_Message_Data_BC_MESSAGE_WORD_02" bit 8
   314: 'BC_MESSAGE_WORD_02_BIT_1', class BC Messages, trigger "64_Message_Data_BC_MESSAGE_WORD_02" bit 9
   315: 'BC_MESSAGE_WORD_02_BIT_2', class BC Messages, trigger "64_Message_Data_BC_MESSAGE_WORD_02" bit 10
   316: 'BC_MESSAGE_WORD_02_BIT_3', class BC Messages, trigger "64_Message_Data_BC_MESSAGE_WORD_02" bit 11
   317: 'BC_MESSAGE_WORD_02_BIT_4', class BC Messages, trigger "64_Message_Data_BC_MESSAGE_WORD_02" bit 12
   318: 'BC_MESSAGE_WORD_02_BIT_5', class BC Messages, trigger "64_Message_Data_BC_MESSAGE_WORD_02" bit 13
   319: 'BC_MESSAGE_WORD_02_BIT_6', class BC Messages, trigger "64_Message_Data_BC_MESSAGE_WORD_02" bit 14
   320: 'BC_MESSAGE_WORD_02_BIT_7', class BC Messages, trigger "64_Message_Data_BC_MESSAGE_WORD_02" bit 15
   321: 'IGG_EVENT_WORD_01_BIT_8', class IGG Events, trigger "66_Event_Data_IGG_EVENT_WORD_01" bit 0
   322: 'IGG_EVENT_WORD_01_BIT_9', class IGG Events, trigger "66_Event_Data_IGG_EVENT_WORD_01" bit 1
   323: 'IGG_EVENT_WORD_01_BIT_10', class IGG Events, trigger "66_Event_Data_IGG_EVENT_WORD_01" bit 2
   324: 'IGG_EVENT_WORD_01_BIT_11', class IGG Events, trigger "66_Event_Data_IGG_EVENT_WORD_01" bit 3
   325: 'IGG_EVENT_WORD_01_BIT_12', class IGG Events, trigger "66_Event_Data_IGG_EVENT_WORD_01" bit 4
   326: 'IGG_EVENT_WORD_01_BIT_13', class IGG Events, trigger "66_Event_Data_IGG_EVENT_WORD_01" bit 5
   327: 'IGG_EVENT_WORD_01_BIT_14', class IGG Events, trigger "66_Event_Data_IGG_EVENT_WORD_01" bit 6
   328: 'IGG_EVENT_WORD_01_BIT_15', class IGG Events, trigger "66_Event_Data_IGG_EVENT_WORD_01" bit 7
   329: 'IGG_EVENT_WORD_01_BIT_0', class IGG Events, trigger "66_Event_Data_IGG_EVENT_WORD_01" bit 8
   330: 'IGG_EVENT_WORD_01_BIT_1', class IGG Events, trigger "66_Event_Data_IGG_EVENT_WORD_01" bit 9
   331: 'IGG_EVENT_WORD_01_BIT_2', class IGG Events, trigger "66_Event_Data_IGG_EVENT_WORD_01" bit 10
   332: 'IGG_EVENT_WORD_01_BIT_3', class IGG Events, trigger "66_Event_Data_IGG_EVENT_WORD_01" bit 11
   333: 'IGG_EVENT_WORD_01_BIT_4', class IGG Events, trigger "66_Event_Data_IGG_EVENT_WORD_01" bit 12
   334: 'IGG_EVENT_WORD_01_BIT_5', class IGG Events, trigger "66_Event_Data_IGG_EVENT_WORD_01" bit 13
   335: 'IGG_EVENT_WORD_01_BIT_6', class IGG Events, trigger "66_Event_Data_IGG_EVENT_WORD_01" bit 14
   336: 'IGG_EVENT_WORD_01_BIT_7', class IGG Events, trigger "66_Event_Data_IGG_EVENT_WORD_01" bit 15
   337: 'IGG_EVENT_WORD_02_BIT_8', class IGG Events, trigger "66_Event_Data_IGG_EVENT_WORD_02" bit 0
   338: 'IGG_EVENT_WORD_02_BIT_9', class IGG Events, trigger "66_Event_Data_IGG_EVENT_WORD_02" bit 1
   339: 'IGG_EVENT_WORD_02_BIT_10', class IGG Events, trigger "66_Event_Data_IGG_EVENT_WORD_02" bit 2
   340: 'IGG_EVENT_WORD_02_BIT_11', class IGG Events, trigger "66_Event_Data_IGG_EVENT_WORD_02" bit 3
   341: 'IGG_EVENT_WORD_02_BIT_12', class IGG Events, trigger "66_Event_Data_IGG_EVENT_WORD_02" bit 4
   342: 'IGG_EVENT_WORD_02_BIT_13', class IGG Events, trigger "66_Event_Data_IGG_EVENT_WORD_02" bit 5
   343: 'IGG_EVENT_WORD_02_BIT_14', class IGG Events, trigger "66_Event_Data_IGG_EVENT_WORD_02" bit 6
   344: 'IGG_EVENT_WORD_02_BIT_15', class IGG Events, trigger "66_Event_Data_IGG_EVENT_WORD_02" bit 7